(* Logix 5000 project; controller PLC_MCC1300_75F1 vendor 1 type 14 code 166 rev 32.11; software revision 32.04; part 70 of 83 *)
(* tags used below, declared in another part *)
   CM_INPUT_Z200_Sync : CM_INPUT_Z200;
   CONST_rgdDestMask : DINT[32];   // Destination Mask
   CONST_tPlant : UDT_PLANT_CONSTANTS;
   GP_TrackingSearchPlate : GP_TrackingSearchPlate;
   GP_TrackingValidateIndex : GP_TrackingValidateIndex;
   M350_M1_DR : AXIS_CIP_DRIVE;
   M350_xReqStopPrevConvForPos : BOOL;
   M350Popup : MAC_Popup_ZC;
   M350Popup_HMW : MAC_Popup_ZC_HMW;
   M350Popup_PlateFreeTimeout : TIMER;
   M350Popup_xDrivePosEnable : BOOL;
   M350Popup_xQualityComing : BOOL;
   TMP_d : DINT;
   TMP_dDiffPhotocellStartConv0 : DINT;
   TMP_dEndSearch0 : DINT;
   TMP_dFixedSideOffset : DINT;
   TMP_dHalfConveyorLength : DINT;
   TMP_dHalfPlateLength : DINT;
   TMP_dIndex : DINT;
   TMP_dStartSearch0 : DINT;
   TMP_xAllLiteToCullet : BOOL;
   TMP_xAtLeastOneForQuality : BOOL;
   TMP_xAtLeastOneForSideLeg : BOOL;
   TMP_xPosHead : BOOL;
   xAlwaysOFF : BOOL;
   xAlwaysON : BOOL;
   xDebugOFF : BOOL;
   Z300_BufferPlate : UDT_LINE_BUFFER_PLATE;
   Z300_Conveyor : UDT_StandConv[29];
   Z300_Conveyor_IN_MOTION : MAC_Conveyor_ZC_IN_MOTION[29];
   Z300_Conveyor_OUT_MOTION : MAC_Conveyor_ZC_OUT_MOTION[29];
   Z300_LineTracking : UDT_LINE_TRACKING;
(* MainProgram, continued *)

ROUTINE M350PopupManagement   (* ladder *)
   // #####_CONSTANTS_#####
   0: NOP();
   1: MOV(CONST_rgdDestMask[29],M350Popup.AUX_dDestMaskOppOpSide)MOV(30000,TMP_dFixedSideOffset)DIV(Z300_LineTracking.rgtTrkConv[21].dLengthConveyor,2,TMP_dHalfConveyorLength);
   // #####_MATCH_#####
   2: NOP();
   3: MOV(Z300_LineTracking.rgtTrkConv[21].dStartPosition_cmm,M350Popup.AUX_dStartPosition_cmm)MOV(Z300_LineTracking.rgtTrkConv[21].dEndPosition_cmm,M350Popup.AUX_dEndPosition_cmm);
   4: SUB(Z300_LineTracking.rgtTrkConv[21].dStartPosition_cmm,20000,M350Popup.AUX_dPosPhotocell_cmm)SUB(Z300_LineTracking.rgtTrkConv[21].dStartPosition_cmm,M350Popup.AUX_dPosPhotocell_cmm,TMP_dDiffPhotocellStartConv0)MOV(50,M350Popup.tmOF_Wait.PRE)[LEQ(CM_INPUT_Z200_Sync.dLehrSpeed_mm_min,17000) MOV(9000,M350Popup.tmON_Saturation.PRE) ,GRT(CM_INPUT_Z200_Sync.dLehrSpeed_mm_min,17000) MOV(9000,M350Popup.tmON_Saturation.PRE) ];
   5: SUB(M350Popup.AUX_dPosPhotocell_cmm,250000,TMP_dStartSearch0)SUB(M350Popup.AUX_dPosPhotocell_cmm,-50000,TMP_dEndSearch0);
   // Set Positioning Type
   6: XIC(xAlwaysON)OTE(TMP_xPosHead);
   // ##### PREVIOUS CONVEYOR #####
   7: NOP();
   // Search plate limits
   8: MUL(M350Popup.AUX_dSpeedConveyor_mm_min,M350Popup.AUX_dReactionTime_ms,TMP_d)DIV(TMP_d,600,M350Popup.AUX_tSearchPlateData.dReaction_cmm);
   9: MOV(TMP_dStartSearch0,M350Popup.AUX_tSearchPlateData.dPositionDecision_cmm)MOV(TMP_dEndSearch0,M350Popup.AUX_tSearchPlateData.dPositionStopSearch_cmm)ADD(Z300_LineTracking.rgtTrkConv[21].dEndPosition_cmm,220000,M350Popup.AUX_tSearchPlateData.dPositionStopHooked_cmm);
   // Search plate on previous conveyor (reverse search)
   10: XIO(M350Popup.AUX_tSearchPlateData.xPlateHooked)GP_TrackingSearchPlate(GP_TrackingSearchPlate,M350Popup.AUX_tSearchPlateData.dPositionStopSearch_cmm,M350Popup.AUX_tSearchPlateData.dPositionDecision_cmm,0,Z300_LineTracking,M350Popup.AUX_tSearchPlateData.tResult,CONST_tPlant.dNumOfConveyors,CONST_tPlant.dNumCapsConveyor,Z300_BufferPlate);
   11: XIO(Z300_LineTracking.rgtTrkConv[20].xGlassPresence)XIO(Z300_LineTracking.rgtTrkConv[21].xGlassPresence)XIC(TMP_xPosHead)XIO(M350Popup.AUX_tSearchPlateData.tResult.xHeadPresence)MOV(0,M350Popup.AUX_tSearchPlateData.dIndex)MOV(0,M350Popup.AUX_dIndexHead);
   12: XIO(Z300_LineTracking.rgtTrkConv[20].xGlassPresence)XIO(Z300_LineTracking.rgtTrkConv[21].xGlassPresence)XIO(TMP_xPosHead)XIO(M350Popup.AUX_tSearchPlateData.tResult.xTailPresence)MOV(0,M350Popup.AUX_tSearchPlateData.dIndex)MOV(0,M350Popup.AUX_dIndexTail);
   13: XIC(TMP_xPosHead)XIC(M350Popup.AUX_tSearchPlateData.tResult.xHeadPresence)MOV(M350Popup.AUX_tSearchPlateData.tResult.rgdHeadPointer[0],M350Popup.AUX_dIndexHead);
   14: XIO(TMP_xPosHead)XIC(M350Popup.AUX_tSearchPlateData.tResult.xTailPresence)MOV(M350Popup.AUX_tSearchPlateData.tResult.rgdTailPointer[0],M350Popup.AUX_dIndexTail);
   15: XIO(M350Popup.AUX_tSearchPlateData.xPlateHooked)[XIC(TMP_xPosHead) XIC(M350Popup.AUX_tSearchPlateData.tResult.xHeadPresence) MOV(M350Popup.AUX_tSearchPlateData.tResult.rgdHeadPointer[0],M350Popup.AUX_tSearchPlateData.dIndex) ,XIO(TMP_xPosHead) XIC(M350Popup.AUX_tSearchPlateData.tResult.xTailPresence) MOV(M350Popup.AUX_tSearchPlateData.tResult.rgdTailPointer[0],M350Popup.AUX_tSearchPlateData.dIndex) ][OSR(M350Popup.AUX_tSearchPlateData.OSR_xPlateInWindows,M350Popup.AUX_tSearchPlateData.OS_xPlateInWindows) ,OSF(M350Popup.AUX_tSearchPlateData.OSF_xPlateInWindows,M350Popup.AUX_tSearchPlateData.OF_xPlateInWindows) ];
   16: GRT(M350Popup.AUX_tSearchPlateData.dIndex,0)[OTU(TMP_xAtLeastOneForSideLeg) ,OTU(TMP_xAtLeastOneForQuality) ,OTL(TMP_xAllLiteToCullet) ];
   // Quality plate redestination for quality table not available
   17: GRT(M350Popup.AUX_tSearchPlateData.dIndex,0)JSR(sbrCheckConvoyZCDestination,5,M350Popup.AUX_tSearchPlateData.dIndex,M350Popup.AUX_dDestMaskOppOpSide,CONST_rgdDestMask[24],TMP_xAtLeastOneForQuality,TMP_xAllLiteToCullet,TMP_xAtLeastOneForQuality,TMP_xAllLiteToCullet)XIC(TMP_xAtLeastOneForQuality)[JSR(sbrRedestConvoyCapZC,5,M350Popup.AUX_tSearchPlateData.dIndex,M350Popup.AUX_dDestMaskOppOpSide,0,1,CONST_rgdDestMask[24]) ,MOV(0,M350Popup.AUX_tSearchPlateData.dIndex) ];
   // Verify destination
   18: GRT(M350Popup.AUX_tSearchPlateData.dIndex,0)[JSR(sbrCheckConvoyZCDestination,5,M350Popup.AUX_tSearchPlateData.dIndex,M350Popup.AUX_dDestMaskOpSide,CONST_rgdDestMask[24],TMP_xAtLeastOneForSideLeg,TMP_xAllLiteToCullet,TMP_xAtLeastOneForSideLeg,TMP_xAllLiteToCullet) XIC(TMP_xAtLeastOneForSideLeg) ,JSR(sbrCheckConvoyZCDestination,5,M350Popup.AUX_tSearchPlateData.dIndex,M350Popup.AUX_dDestMaskOppOpSide,CONST_rgdDestMask[24],TMP_xAtLeastOneForQuality,TMP_xAllLiteToCullet,TMP_xAtLeastOneForQuality,TMP_xAllLiteToCullet) XIC(TMP_xAtLeastOneForQuality) ][OTE(M350Popup.ST_xPlateComingToPopup) ,XIO(TMP_xAtLeastOneForSideLeg) XIO(TMP_xAtLeastOneForQuality) MOV(M350Popup.AUX_tSearchPlateData.dIndex,M350Popup.AUX_dIndexPlateFree) ];
   19: XIO(Z300_LineTracking.rgtTrkConv[20].xGlassPresence)XIO(Z300_LineTracking.rgtTrkConv[21].xGlassPresence)MOV(0,M350Popup.AUX_dIndexPlateFree);
   20: GP_TrackingValidateIndex(GP_TrackingValidateIndex,Z300_BufferPlate,M350Popup.AUX_tSearchPlateData.dIDMemory,M350Popup.AUX_tSearchPlateData.dIndex,M350Popup.AUX_tSearchPlateData.xIndexCons);
   // Check plate dimension
   21: XIC(M350Popup.ST_xPlateComingToPopup)MOV(M350Popup.AUX_tSearchPlateData.dIndex,TMP_dIndex)[LEQ(Z300_BufferPlate.rgtPlate[TMP_dIndex].tData.dTotalCaps,1) GEQ(Z300_BufferPlate.rgtPlate[TMP_dIndex].tData.dLength_cmm,CONST_tPlant.rgdLiteLimits_cmm[6]) OTE(M350Popup.ST_xPlateToSingleComing) ,GRT(Z300_BufferPlate.rgtPlate[TMP_dIndex].tData.dTotalCaps,1) [LEQ(Z300_BufferPlate.rgtPlate[TMP_dIndex].tData.dLength_cmm,CONST_tPlant.rgdConvoyLimits_cmm[2]) ,XIO(xDebugOFF) ] OTE(M350Popup.ST_xConvoyComing) ];
   22: [XIC(Z300_Conveyor[20].xReqStop) ,XIO(xAlwaysOFF) ]XIC(M350Popup.ST_xPhasesInProgress)XIO(M350Popup.PH_xDescend)TOF(M350Popup.tmOF_Wait,?,?);
   // Plate has left popup conveyors
   23: GRT(M350Popup.AUX_dIndexPlateFree,0)MOV(M350Popup.AUX_dIndexPlateFree,TMP_dIndex)GEQ(Z300_BufferPlate.rgtPlate[TMP_dIndex].tTracking.dPositionTail_cmm,M350Popup.AUX_dEndPosition_cmm)MOV(0,M350Popup.AUX_dIndexPlateFree);
   // Stop previuos conveyor if no condition on pop-up conveyor
   24: [[XIC(M350Popup.ST_xPlateToSingleComing) ,XIC(M350Popup.ST_xConvoyComing) ] [XIO(M350Popup.ST_xInitialConditionForRise) ,XIC(Z300_LineTracking.rgtTrkConv[21].xGlassPresence) ,XIC(M350Popup.ST_xPlateUnderPopup) EQU(M350Popup.AUX_dIndexPositioning,0) ] ,XIC(M350_xReqStopPrevConvForPos) ,XIC(Z300_Conveyor[21].xReqExtStopLoadNewPlate) ,XIC(M350Popup.ST_xPlateInPositionToRise) ,XIO(M350Popup.INPUT_xPopupLow) XIO(M350Popup.PH_xDescend) ,XIC(M350Popup.ST_xPhasesInProgress) XIO(M350Popup.PH_xDescend) ,XIC(M350Popup.tmOF_Wait.DN) XIO(M350Popup.PH_xDescend) ,XIC(Z300_Conveyor[21].ST_xCleaningEnabled) XIO(Z300_Conveyor[20].ST_xCleaningEnabled) ,GRT(M350Popup.AUX_dIndexPositioning,0) [GRT(M350Popup.AUX_tSearchPlateData.dIndex,0) NEQ(M350Popup.AUX_tSearchPlateData.dIndex,M350Popup.AUX_dIndexPositioning) ,GRT(M350Popup.AUX_dIndexPlatePositioned,0) NEQ(M350Popup.AUX_dIndexPlatePositioned,M350Popup.AUX_dIndexPositioning) ] ,GRT(M350Popup.AUX_dIndexPlateFree,0) MOV(M350Popup.AUX_dIndexPlateFree,TMP_dIndex) [XIC(M350Popup.ST_xPlateToSingleComing) [XIC(Z300_Conveyor[21].ST_xRotationFeedback) SUB(M350Popup.AUX_dEndPosition_cmm,Z300_Conveyor[21].AUX_rgdDecSpace_cmm[0],TMP_d) ,XIO(Z300_Conveyor[21].ST_xRotationFeedback) MOV(M350Popup.AUX_dEndPosition_cmm,TMP_d) ] LES(Z300_BufferPlate.rgtPlate[TMP_dIndex].tTracking.dPositionTail_cmm,TMP_d) ,[XIC(M350Popup.ST_xPlateToBothComing) ,XIC(M350Popup.ST_xConvoyComing) ] [XIC(Z300_Conveyor[21].ST_xRotationFeedback) SUB(M350Popup.AUX_dEndPosition_cmm,Z300_Conveyor[21].AUX_rgdDecSpace_cmm[0],TMP_d) ,XIO(Z300_Conveyor[21].ST_xRotationFeedback) MOV(M350Popup.AUX_dEndPosition_cmm,TMP_d) ] LES(Z300_BufferPlate.rgtPlate[TMP_dIndex].tTracking.dPositionTail_cmm,TMP_d) ] ]OTE(M350Popup.ST_xConditionToStopPrevious);
   25: XIO(xDebugOFF)XIO(Z300_LineTracking.rgtTrkConv[21].xGlassPresence)XIC(Z300_Conveyor[21].ST_xRotationFeedback)[GRT(M350Popup.AUX_dIndexPlateFree,0) ,GRT(M350Popup.AUX_dIndexPlatePositioned,0) ]MOV(5000,M350Popup_PlateFreeTimeout.PRE)[TON(M350Popup_PlateFreeTimeout,?,?) ,XIC(M350Popup_PlateFreeTimeout.DN) [MOV(0,M350Popup.AUX_dIndexPlateFree) ,MOV(0,M350Popup.AUX_dIndexPlatePositioned) ] ];
   26: XIC(M350Popup.ST_xConditionToStopPrevious)[XIC(xAlwaysOFF) XIC(Z300_LineTracking.rgtTrkConv[20].xGlassPresCom) GRT(Z300_LineTracking.rgtTrkConv[20].dHeadPosition_cmm,0) ,XIO(xDebugOFF) SUB(Z300_Conveyor[20].AUX_rgdLoadPreset_cmm[0],0,TMP_d) GEQ(Z300_LineTracking.rgtTrkConv[20].dHeadPosition_cmm,TMP_d) ,XIC(xDebugOFF) SUB(Z300_Conveyor[20].AUX_rgdLoadPresetWithRestart_cmm[0],10000,TMP_d) GEQ(Z300_LineTracking.rgtTrkConv[20].dHeadPosition_cmm,TMP_d) ][XIO(Z300_LineTracking.rgtTrkConv[20].xPlatePassageNext) ,XIO(xAlwaysOFF) ][XIO(Z300_Conveyor[21].OUTPUT_xPositioning.0) XIO(M350Popup.tmON_Positioning.EN) ,[XIC(M350_xReqStopPrevConvForPos) ,XIC(Z300_Conveyor[21].xReqExtStopLoadNewPlate) ] ]OTE(M350Popup.ST_xStopPreviousConveyor);
   // STOP CONVEYOR M322
   27: XIC(M350Popup.ST_xStopPreviousConveyor)OTE(Z300_Conveyor[20].xReqStop);
   28: XIO(xDebugOFF)XIO(Z300_Conveyor[20].xReqStop)[XIO(Z300_LineTracking.rgtTrkConv[21].xGlassPresence) XIO(Z300_LineTracking.rgtTrkConv[22].xGlassPresence) XIC(Z300_Conveyor[21].ST_xRotationFeedback) XIC(Z300_Conveyor[22].ST_xRotationFeedback) XIC(M350Popup.INPUT_xPopupLow) ,XIO(Z300_LineTracking.rgtTrkConv[20].xPlatePassageNext) XIO(Z300_LineTracking.rgtTrkConv[21].xPlatePassagePrevious) XIC(Z300_Conveyor[21].ST_xRotationFeedback) ]OTE(Z300_Conveyor[20].xReqBypassEndStop);
   // #####_POSITIONING_#####
   29: NOP();
   // Hook plate for positioning
   30: XIO(M350Popup.ST_xPlatePresentOnPopup)XIO(M350Popup.ST_xPlatePresence)XIO(M350Popup.AUX_tSearchPlateData.xPlateHooked)EQU(M350Popup.AUX_dIndexPositioning,0)GRT(M350Popup.AUX_tSearchPlateData.dIndex,0)XIC(M350Popup.AUX_tSearchPlateData.xIndexCons)MOV(M350Popup.AUX_tSearchPlateData.dIndex,TMP_dIndex)GRT(Z300_BufferPlate.rgtPlate[TMP_dIndex].tTracking.dPositionHead_cmm,M350Popup.AUX_tSearchPlateData.dPositionDecision_cmm)XIC(M350Popup.ST_xPlateComingToPopup)XIO(Z300_LineTracking.rgtTrkConv[21].xGlassPresence)XIO(Z300_Conveyor[21].OUTPUT_xPositioning.0)XIO(M350Popup.ST_xPlateInPositionToRise)[OTL(M350Popup.AUX_tSearchPlateData.xPlateHooked) ,MOV(M350Popup.AUX_tSearchPlateData.dIndex,M350Popup.AUX_dIndexPositioning) ,JSR(sbrTrackingPositioningStart,2,M350Popup.AUX_dIndexPositioning,TMP_xPosHead) ,GRT(M350Popup.tSearchPlateStop.rgdHeadPointer[0],0) MOV(M350Popup.tSearchPlateStop.rgdHeadPointer[0],M350Popup.AUX_dIndexPlateFree) ,XIC(TMP_xAtLeastOneForQuality) OTL(M350Popup_xQualityComing) ];
   31: GP_TrackingValidateIndex(GP_TrackingValidateIndex,Z300_BufferPlate,M350Popup.AUX_dMemoryPositioning,M350Popup.AUX_dIndexPositioning,M350Popup.ST_xIndexConsPositioning);
   // Check plate dimension
   32: XIC(M350Popup.AUX_tSearchPlateData.xPlateHooked)XIC(M350Popup.ST_xIndexConsPositioning)XIO(M350Popup.ST_xPlateToSinglePositioning)XIO(M350Popup.ST_xConvoyPositioning)MOV(M350Popup.AUX_dIndexPositioning,TMP_dIndex)[LEQ(Z300_BufferPlate.rgtPlate[TMP_dIndex].tData.dTotalCaps,1) GEQ(Z300_BufferPlate.rgtPlate[TMP_dIndex].tData.dLength_cmm,CONST_tPlant.rgdLiteLimits_cmm[6]) OTL(M350Popup.ST_xPlateToSinglePositioning) ,GRT(Z300_BufferPlate.rgtPlate[TMP_dIndex].tData.dTotalCaps,1) LEQ(Z300_BufferPlate.rgtPlate[TMP_dIndex].tData.dLength_cmm,CONST_tPlant.rgdConvoyLimits_cmm[2]) OTL(M350Popup.ST_xConvoyPositioning) ];
   // Positioning request (In case of head positioning also previous conveyors are involved)
   33: XIC(M350Popup.AUX_tSearchPlateData.xPlateHooked)[XIC(M350Popup.ST_xIndexConsPositioning) ,XIO(xDebugOFF) ][XIC(M350Popup.ST_xPlateToSinglePositioning) ,XIC(M350Popup.ST_xConvoyPositioning) ]XIO(M350Popup.ST_xPlatePresence)[XIO(M350Popup.ST_xPlateUnderPopup) ,XIO(xAlwaysOFF) ]XIO(Z300_LineTracking.rgtTrkConv[21].xGlassPresence)XIO(Z300_Conveyor[21].xReqStop)XIC(M350Popup.ST_xOutputEnable)[XIC(M350Popup.INPUT_xPopupLow) XIC(M350Popup.ST_xInitialConditionForRise) ,XIC(M350Popup.OUTPUT_xPopupDescent) ]XIO(Z300_Conveyor[21].xReqPositioningHead)XIO(Z300_Conveyor[21].xReqPositioningTail)TON(M350Popup.tmON_Positioning,?,?)XIC(M350Popup.tmON_Positioning.DN)[XIC(TMP_xPosHead) OTL(Z300_Conveyor[21].xReqPositioningHead) ,XIO(TMP_xPosHead) OTL(Z300_Conveyor[21].xReqPositioningTail) ,OTE(M350Popup.OS_xStartPositioning) ,OTU(Z300_Conveyor_OUT_MOTION[21].DR_MAR_M[0].PC) ,OTU(Z300_Conveyor_IN_MOTION[21].DR_MAR_M[0].PC) ,OTU(Z300_Conveyor_OUT_MOTION[21].DR_MAM_M[0].PC) ,OTU(Z300_Conveyor_IN_MOTION[21].DR_MAM_M[0].PC) ];
   34: DIV(360000,2,TMP_dHalfConveyorLength);
   // Target calculation
   35: XIC(M350Popup.OS_xStartPositioning)[XIC(M350Popup.ST_xIndexConsPositioning) ,XIO(xDebugOFF) ]MOV(M350Popup.AUX_tSearchPlateData.dIndex,TMP_dIndex)[XIC(M350Popup.ST_xPlateToSinglePositioning) ADD(TMP_dDiffPhotocellStartConv0,TMP_dFixedSideOffset,TMP_d) [XIC(TMP_xPosHead) [XIO(Z300_BufferPlate.rgtPlate[TMP_dIndex].tData.rgtCap[0].rgxRequest.1) ADD(TMP_d,Z300_BufferPlate.rgtPlate[TMP_dIndex].tData.dLength_cmm,M350Popup.AUX_dReqTarget_cmm) ,XIC(Z300_BufferPlate.rgtPlate[TMP_dIndex].tData.rgtCap[0].rgxRequest.1) ADD(TMP_d,300000,M350Popup.AUX_dReqTarget_cmm) ] ,XIO(TMP_xPosHead) MOV(TMP_d,M350Popup.AUX_dReqTarget_cmm) ] ,XIC(M350Popup.ST_xConvoyPositioning) DIV(Z300_BufferPlate.rgtPlate[TMP_dIndex].tData.rgtCap[0].dConvTotLength_cmm,2,TMP_dHalfPlateLength) ADD(TMP_dDiffPhotocellStartConv0,TMP_dHalfConveyorLength,TMP_d) [XIC(TMP_xPosHead) ADD(TMP_d,TMP_dHalfPlateLength,M350Popup.AUX_dReqTarget_cmm) ,XIO(TMP_xPosHead) SUB(TMP_d,TMP_dHalfPlateLength,M350Popup.AUX_dReqTarget_cmm) ] ,XIC(M350Popup_xQualityComing) ADD(TMP_dDiffPhotocellStartConv0,325000,TMP_d) [XIC(TMP_xPosHead) ,XIO(TMP_xPosHead) SUB(TMP_d,Z300_BufferPlate.rgtPlate[TMP_dIndex].tData.dLength_cmm,TMP_d) ] MOV(TMP_d,M350Popup.AUX_dReqTarget_cmm) ];
   // Final drive target (In case of head positioning also previous conveyors are involved)
   36: XIC(M350Popup.OS_xStartPositioning)[XIC(M350Popup.ST_xIndexConsPositioning) ,XIO(xDebugOFF) ]SUB(M350Popup.AUX_dReqTarget_cmm,TMP_dDiffPhotocellStartConv0,TMP_d)ADD(TMP_d,Z300_LineTracking.rgtTrkConv[21].dStartPosition_cmm,TMP_d)ADD(TMP_d,220000,M350Popup.AUX_dPosTimeout)[XIC(M350Popup.ST_xPlateToSinglePositioning) ADD(M350Popup.AUX_dReqTarget_cmm,M350Popup_HMW.dSingleCapOffset_cmm,Z300_Conveyor[21].AUX_rgdTarget_cmm[0]) ,XIC(M350Popup.ST_xConvoyPositioning) ADD(M350Popup.AUX_dReqTarget_cmm,M350Popup_HMW.dConvoyOffset_cmm,Z300_Conveyor[21].AUX_rgdTarget_cmm[0]) ,XIC(M350Popup_xQualityComing) MOV(M350Popup.AUX_dReqTarget_cmm,Z300_Conveyor[21].AUX_rgdTarget_cmm[0]) ]XIC(TMP_xPosHead)[MOV(Z300_Conveyor[21].AUX_rgdTarget_cmm[0],Z300_Conveyor[20].AUX_rgdTarget_cmm[0]) ,MOV(Z300_Conveyor[21].AUX_rgdTarget_cmm[0],Z300_Conveyor[20].AUX_rgdTarget_cmm[1]) ];
   37: XIC(Z300_LineTracking.rgtTrkConv[21].xGlassPresence)MOV(M350Popup.AUX_dIndexPositioning,TMP_dIndex)GRT(TMP_dIndex,0)LES(Z300_BufferPlate.rgtPlate[TMP_dIndex].tData.dTotalCaps,2)[XIC(Z300_Conveyor[21].OUTPUT_xPositioning.0) GEQ(Z300_BufferPlate.rgtPlate[TMP_dIndex].tTracking.dPositionHead_cmm,M350Popup.AUX_dStartPosition_cmm) XIC(M350Popup_xDrivePosEnable) XIO(M350_M1_DR.Registration1InputStatus) ,XIC(Z300_Conveyor[21].xReqExtStopLoadNewPlate) ]OTE(Z300_Conveyor[21].xReqExtStopLoadNewPlate);
   38: XIC(Z300_Conveyor[21].OUTPUT_xPositioning.0)[XIC(Z300_Conveyor_IN_MOTION[21].DR_MAM_M[0].PC) ,XIC(xAlwaysOFF) ADD(Z300_LineTracking.rgtTrkConv[21].dStartPosition_cmm,Z300_Conveyor[21].AUX_rgdTarget_cmm[0],TMP_d) SUB(TMP_d,Z300_LineTracking.rgtTrkConv[21].dActualRamp_cmm[0],TMP_d) GEQ(Z300_BufferPlate.rgtPlate[TMP_dIndex].tTracking.dPositionHead_cmm,TMP_d) ][OTE(Z300_Conveyor[21].ST_xPositionReached) ,MOV(M350Popup.AUX_dIndexPositioning,TMP_dIndex) JSR(sbrTrackingPositioningDone,3,TMP_dIndex,TMP_xPosHead,Z300_Conveyor[21].AUX_rgdTarget_cmm[0]) ];
   // Head positioning done
   39: XIC(Z300_Conveyor[21].xReqPositioningHead)[XIC(Z300_Conveyor[21].ST_xPositionReached) ,XIC(M350Popup.OS_xTimeoutPositioning) ,XIC(xDebugOFF) XIO(M350Popup.ST_xIndexConsPositioning) ,XIC(Z300_Conveyor[21].ST_xFaulted) ][OTU(Z300_Conveyor[21].xReqPositioningHead) ,OTU(Z300_Conveyor[20].xReqPositioningHead) ,XIO(Z300_Conveyor[21].ST_xFaulted) XIO(M350Popup.OS_xTimeoutPositioning) XIC(M350Popup.ST_xIndexConsPositioning) MOV(M350Popup.AUX_dIndexPositioning,TMP_dIndex) [OTL(Z300_BufferPlate.rgtPlate[TMP_dIndex].tData.tFlag.tConveyor.xDoneHeadPositioning) ,JSR(sbrTrackingPositioningDone,3,TMP_dIndex,TMP_xPosHead,Z300_Conveyor[21].AUX_rgdTarget_cmm[0]) ,MOV(M350Popup.AUX_dIndexPositioning,M350Popup.AUX_dIndexPlatePositioned) ] ,MOV(0,M350Popup.AUX_dIndexHead) ];
   // When plate tail has passed previous conveyor remove positioning
   40: XIC(Z300_Conveyor[20].xReqPositioningHead)[XIO(M350Popup.ST_xPrevConvFreeAfterPos) NEQ(M350Popup.AUX_dIndexPositioning,0) ,XIC(M350Popup.ST_xPrevConvFreeAfterPos) EQU(M350Popup.AUX_dIndexPositioning,M350Popup.AUX_dLastIndexFreeForPos) ][XIC(Z300_Conveyor[20].xReqPositioningHead) MOV(M350Popup.AUX_dIndexPositioning,TMP_dIndex) GEQ(Z300_BufferPlate.rgtPlate[TMP_dIndex].tTracking.dPositionTail_cmm,Z300_LineTracking.rgtTrkConv[20].dEndPosition_cmm) ,XIC(M350Popup.ST_xPrevConvFreeAfterPos) ][OTU(Z300_Conveyor[20].xReqPositioningHead) ,OTE(M350Popup.ST_xPrevConvFreeAfterPos) ,ONS(M350Popup.OS_xLastFreeForPos) MOV(M350Popup.AUX_dIndexPositioning,M350Popup.AUX_dLastIndexFreeForPos) ];
   // Tail positioning done
   41: XIC(Z300_Conveyor[21].xReqPositioningTail)[XIC(Z300_Conveyor[21].ST_xPositionReached) ,XIC(M350Popup.OS_xTimeoutPositioning) ,XIO(M350Popup.ST_xIndexConsPositioning) ,XIC(Z300_Conveyor[21].ST_xFaulted) ][OTU(Z300_Conveyor[21].xReqPositioningTail) ,XIO(Z300_Conveyor[21].ST_xFaulted) XIO(M350Popup.OS_xTimeoutPositioning) MOV(M350Popup.AUX_tSearchPlateData.dIndex,TMP_dIndex) [OTL(Z300_BufferPlate.rgtPlate[TMP_dIndex].tData.tFlag.tConveyor.xDoneTailPositioning) ,JSR(sbrTrackingPositioningDone,3,TMP_dIndex,TMP_xPosHead,Z300_Conveyor[21].AUX_rgdTarget_cmm[0]) ,MOV(M350Popup.AUX_dIndexPositioning,M350Popup.AUX_dIndexPlatePositioned) ] ,MOV(0,M350Popup.AUX_dIndexTail) ];
   // Timeout positioning
   42: [XIC(Z300_Conveyor[21].xReqPositioningHead) MOV(M350Popup.AUX_dIndexPositioning,TMP_dIndex) GEQ(Z300_BufferPlate.rgtPlate[TMP_dIndex].tTracking.dPositionHead_cmm,M350Popup.AUX_dPosTimeout) XIO(Z300_BufferPlate.rgtPlate[TMP_dIndex].tData.tFlag.tConveyor.xDoneHeadPositioning) ,XIC(Z300_Conveyor[21].xReqPositioningTail) MOV(M350Popup.AUX_dIndexPositioning,TMP_dIndex) GEQ(Z300_BufferPlate.rgtPlate[TMP_dIndex].tTracking.dPositionTail_cmm,M350Popup.AUX_dPosTimeout) XIO(Z300_BufferPlate.rgtPlate[TMP_dIndex].tData.tFlag.tConveyor.xDoneTailPositioning) ]OTE(M350Popup.OS_xTimeoutPositioning);
   43: XIC(Z300_Conveyor[21].xReqPositioningHead)XIO(M350Popup.AUX_tSearchPlateData.xPlateHooked)OTU(Z300_Conveyor[21].xReqPositioningHead);
   44: XIC(Z300_Conveyor[21].xReqPositioningTail)XIO(M350Popup.AUX_tSearchPlateData.xPlateHooked)OTU(Z300_Conveyor[21].xReqPositioningTail);
   45: XIC(Z300_Conveyor[20].xReqPositioningHead)XIO(M350Popup.AUX_tSearchPlateData.xPlateHooked)OTU(Z300_Conveyor[20].xReqPositioningHead);
   46: XIC(Z300_Conveyor[20].xReqPositioningTail)XIO(M350Popup.AUX_tSearchPlateData.xPlateHooked)OTU(Z300_Conveyor[20].xReqPositioningTail);
